// TIA Portal project "Mes_Con" (V17) (continued)
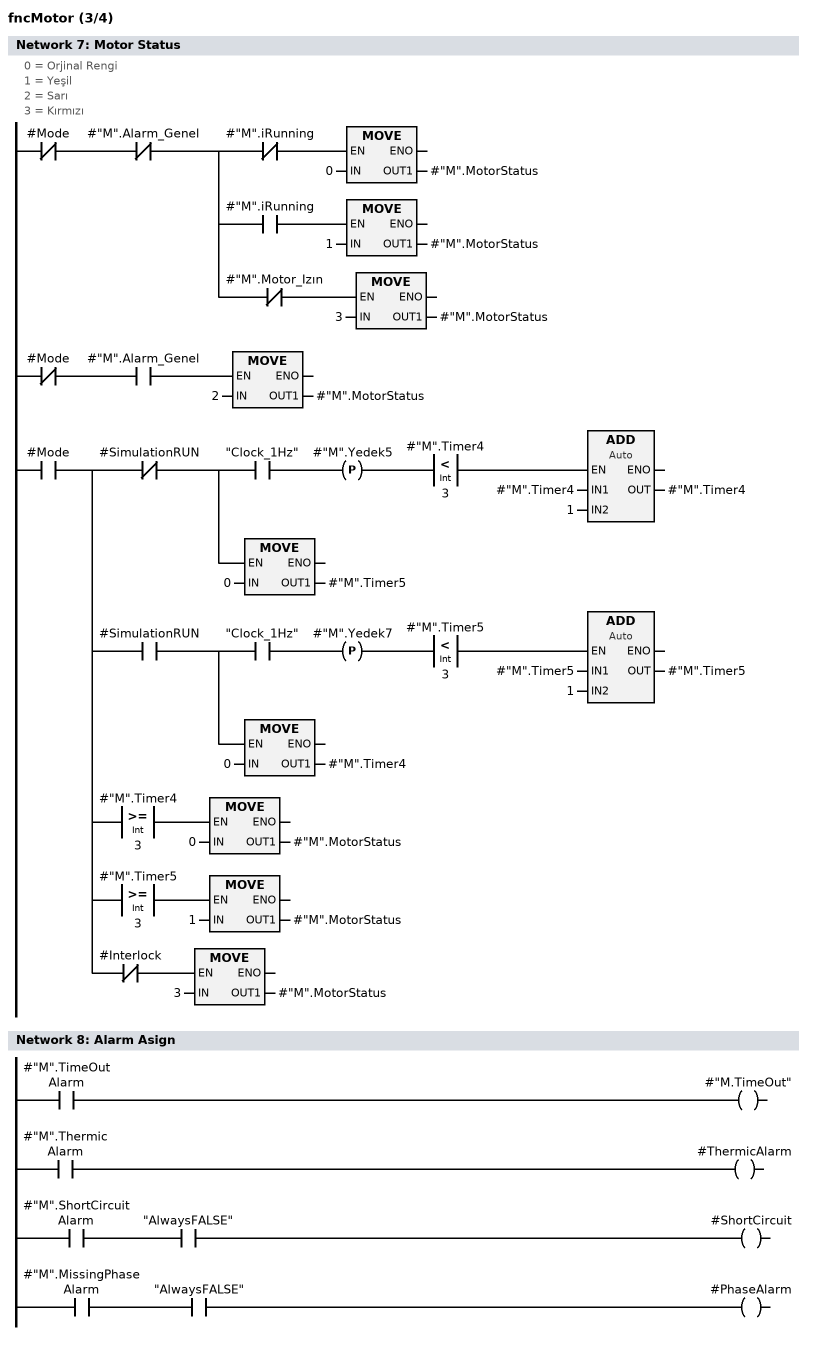
   RUNG wire#powerrail
      I_Contact( #Mode )
      I_Contact( #"M".Alarm_Genel )
      wire#w1
      I_Contact( #"M".iRunning )
      Move(in := 0, out1 => #"M".MotorStatus)
   END_RUNG
   RUNG wire#w1
      Contact( #"M".iRunning )
      Move(in := 1, out1 => #"M".MotorStatus)
   END_RUNG
   RUNG wire#w1
      I_Contact( #"M".Motor_Izın )
      Move(in := 3, out1 => #"M".MotorStatus)
   END_RUNG
   RUNG wire#powerrail
      I_Contact( #Mode )
      Contact( #"M".Alarm_Genel )
      Move(in := 2, out1 => #"M".MotorStatus)
   END_RUNG
   RUNG wire#powerrail
      Contact( #Mode )
      wire#w2
      I_Contact( #SimulationRUN )
      wire#w3
      Contact( "Clock_1Hz" )
      P_Trig( #"M".Yedek5 )
      { S7_Templates := "SrcType := Int" } LT_Contact(in1 := #"M".Timer4, in2 := 3)
      Add(in1 := #"M".Timer4, in2 := 1, out => #"M".Timer4)
   END_RUNG
   RUNG wire#w3
      Move(in := 0, out1 => #"M".Timer5)
   END_RUNG
   RUNG wire#w2
      Contact( #SimulationRUN )
      wire#w4
      Contact( "Clock_1Hz" )
      P_Trig( #"M".Yedek7 )
      { S7_Templates := "SrcType := Int" } LT_Contact(in1 := #"M".Timer5, in2 := 3)
      Add(in1 := #"M".Timer5, in2 := 1, out => #"M".Timer5)
   END_RUNG
   RUNG wire#w4
      Move(in := 0, out1 => #"M".Timer4)
   END_RUNG
   RUNG wire#w2
      { S7_Templates := "SrcType := Int" } GE_Contact(in1 := #"M".Timer4, in2 := 3)
      Move(in := 0, out1 => #"M".MotorStatus)
   END_RUNG
   RUNG wire#w2
      { S7_Templates := "SrcType := Int" } GE_Contact(in1 := #"M".Timer5, in2 := 3)
      Move(in := 1, out1 => #"M".MotorStatus)
   END_RUNG
   RUNG wire#w2
      I_Contact( #Interlock )
      Move(in := 3, out1 => #"M".MotorStatus)
   END_RUNG
   // the same network as SCL:
   #_w1 := NOT #Mode AND NOT #"M".Alarm_Genel;
   IF #_w1 AND NOT #"M".iRunning THEN #"M".MotorStatus := 0; END_IF;
   IF #_w1 AND #"M".iRunning THEN #"M".MotorStatus := 1; END_IF;
   IF #_w1 AND NOT #"M".Motor_Izın THEN #"M".MotorStatus := 3; END_IF;
   IF NOT #Mode AND #"M".Alarm_Genel THEN #"M".MotorStatus := 2; END_IF;
   #_w2 := #Mode AND NOT #SimulationRUN;
   #_w3 := #_w2 AND "Clock_1Hz";
   #_w4 := #_w3 AND NOT #"M".Yedek5;   // rising edge
   #"M".Yedek5 := #_w3;
   IF #_w4 AND (#"M".Timer4 < 3) THEN #"M".Timer4 := #"M".Timer4 + 1; END_IF;
   IF #_w2 THEN #"M".Timer5 := 0; END_IF;
   #_w5 := #Mode AND #SimulationRUN;
   #_w6 := #_w5 AND "Clock_1Hz";
   #_w7 := #_w6 AND NOT #"M".Yedek7;   // rising edge
   #"M".Yedek7 := #_w6;
   IF #_w7 AND (#"M".Timer5 < 3) THEN #"M".Timer5 := #"M".Timer5 + 1; END_IF;
   IF #_w5 THEN #"M".Timer4 := 0; END_IF;
   IF #Mode AND (#"M".Timer4 >= 3) THEN #"M".MotorStatus := 0; END_IF;
   IF #Mode AND (#"M".Timer5 >= 3) THEN #"M".MotorStatus := 1; END_IF;
   IF #Mode AND NOT #Interlock THEN #"M".MotorStatus := 3; END_IF;
END_REGION

REGION Network 8: Alarm Asign
   RUNG wire#powerrail
      Contact( #"M".TimeOutAlarm )
      Coil( #"M.TimeOut" )
   END_RUNG
   RUNG wire#powerrail
      Contact( #"M".ThermicAlarm )
      Coil( #ThermicAlarm )
   END_RUNG
   RUNG wire#powerrail
      Contact( #"M".ShortCircuitAlarm )
      Contact( "AlwaysFALSE" )
      Coil( #ShortCircuit )
   END_RUNG
   RUNG wire#powerrail
      Contact( #"M".MissingPhaseAlarm )
      Contact( "AlwaysFALSE" )
      Coil( #PhaseAlarm )
   END_RUNG
   // the same network as SCL:
   #"M.TimeOut" := #"M".TimeOutAlarm;
   #ThermicAlarm := #"M".ThermicAlarm;
   #ShortCircuit := #"M".ShortCircuitAlarm AND "AlwaysFALSE";
   #PhaseAlarm := #"M".MissingPhaseAlarm AND "AlwaysFALSE";
END_REGION

REGION Network 9: POPUP KAPATMA
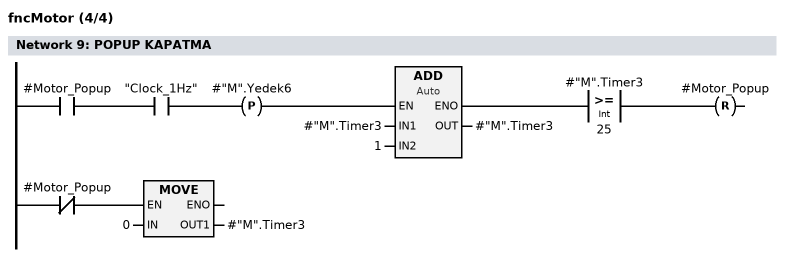
   RUNG wire#powerrail
      Contact( #Motor_Popup )
      Contact( "Clock_1Hz" )
      P_Trig( #"M".Yedek6 )
      Add(in1 := #"M".Timer3, in2 := 1, out => #"M".Timer3)
      { S7_Templates := "SrcType := Int" } GE_Contact(in1 := #"M".Timer3, in2 := 25)
      R_Coil( #Motor_Popup )
   END_RUNG
   RUNG wire#powerrail
      I_Contact( #Motor_Popup )
      Move(in := 0, out1 => #"M".Timer3)
   END_RUNG
   // the same network as SCL:
   #_w1 := #Motor_Popup AND "Clock_1Hz";
   #_w2 := #_w1 AND NOT #"M".Yedek6;   // rising edge
   #"M".Yedek6 := #_w1;
   IF #_w2 THEN #"M".Timer3 := #"M".Timer3 + 1; END_IF;
   IF #_w2 AND (#"M".Timer3 >= 25) THEN #Motor_Popup := FALSE; END_IF;
   IF NOT #Motor_Popup THEN #"M".Timer3 := 0; END_IF;
END_REGION
END_FUNCTION

// folder: Eqp/Valve

FUNCTION "fncValve" : Void   // FC3, LAD
{ S7_Optimized_Access := 'TRUE' }
VERSION : 0.1
   VAR_INPUT
      Mode : Bool;   // 0 = RunTime , 1 = Simulation
      Valve_Opened : Bool;
      Valve_Closed : Bool;
      Interlock : Bool;
   END_VAR
   VAR_OUTPUT
      Valve_Run : Bool;
      Valve_Alarm : Bool;
      Not_Opened : Bool;
      Not_Closed : Bool;
      Not_Signal : Bool;
      Two_Signal : Bool;
   END_VAR
   VAR_IN_OUT
      V : "Valve";
      Vana_Popup : Bool;
   END_VAR
   VAR_TEMP
      SimOpen : Bool;
      SimClose : Bool;
   END_VAR
   VAR_TEMP   // added for the SCL form of the ladder/FBD networks
      _w1 : Bool;
      _w2 : Bool;
      _w3 : Bool;
      _w4 : Bool;
      _w5 : Bool;
      _w6 : Bool;
      _w7 : Bool;
      _w8 : Bool;
      _w9 : Bool;
      _w10 : Bool;
      _w11 : Bool;
      _w12 : Bool;
   END_VAR
BEGIN

REGION Network 1: ATAMA
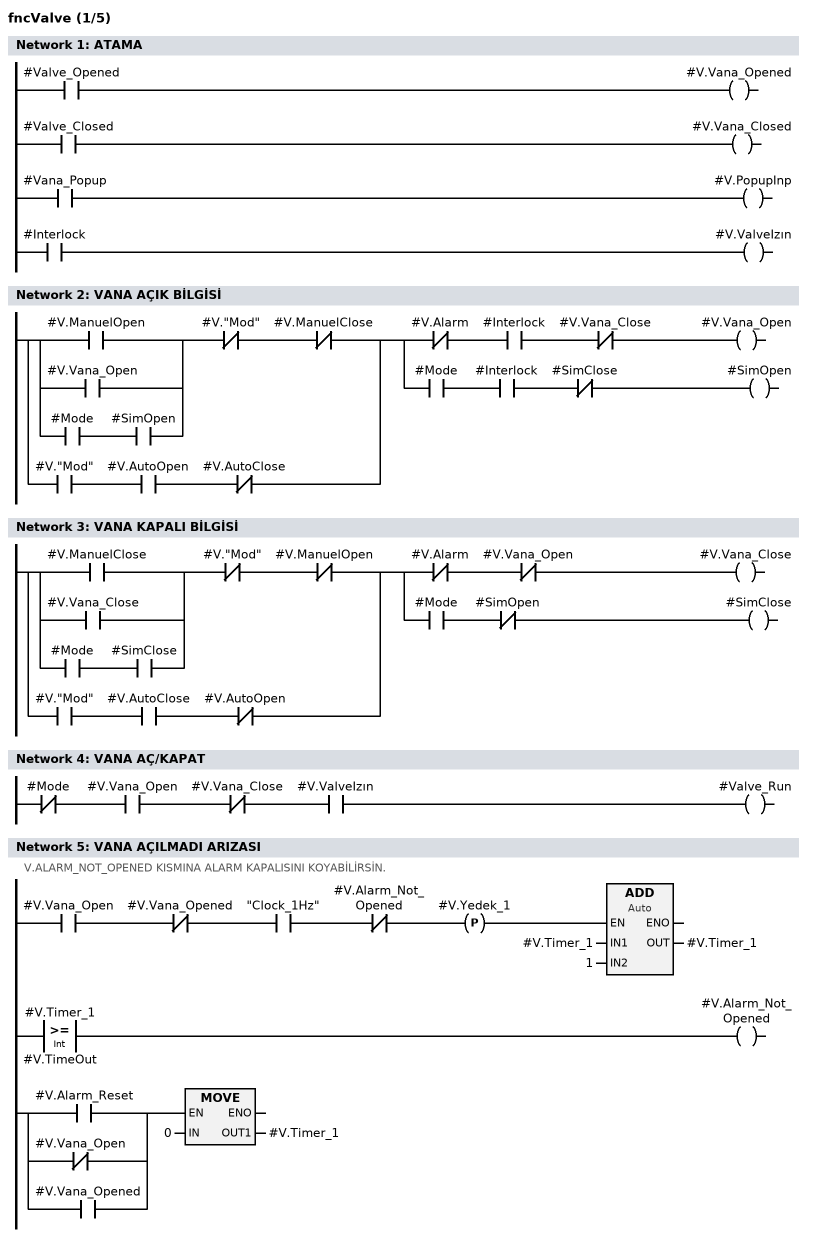
   RUNG wire#powerrail
      Contact( #Valve_Opened )
      Coil( #V.Vana_Opened )
   END_RUNG
   RUNG wire#powerrail
      Contact( #Valve_Closed )
      Coil( #V.Vana_Closed )
   END_RUNG
   RUNG wire#powerrail
      Contact( #Vana_Popup )
      Coil( #V.PopupInp )
   END_RUNG
   RUNG wire#powerrail
      Contact( #Interlock )
      Coil( #V.ValveIzın )
   END_RUNG
   // the same network as SCL:
   #V.Vana_Opened := #Valve_Opened;
   #V.Vana_Closed := #Valve_Closed;
   #V.PopupInp := #Vana_Popup;
   #V.ValveIzın := #Interlock;
END_REGION

REGION Network 2: VANA AÇIK BİLGİSİ
   RUNG wire#powerrail
      Contact( #V.ManuelOpen )
      wire#w1
      I_Contact( #V."Mod" )
      I_Contact( #V.ManuelClose )
      wire#w2
      I_Contact( #V.Alarm )
      Contact( #Interlock )
      I_Contact( #V.Vana_Close )
      Coil( #V.Vana_Open )
   END_RUNG
   RUNG wire#powerrail
      Contact( #V.Vana_Open )
   END_RUNG wire#w1
   RUNG wire#powerrail
      Contact( #Mode )
      Contact( #SimOpen )
   END_RUNG wire#w1
   RUNG wire#powerrail
      Contact( #V."Mod" )
      Contact( #V.AutoOpen )
      I_Contact( #V.AutoClose )
   END_RUNG wire#w2
   RUNG wire#w2
      Contact( #Mode )
      Contact( #Interlock )
      I_Contact( #SimClose )
      Coil( #SimOpen )
   END_RUNG
   // the same network as SCL:
   #_w1 := ((#V.ManuelOpen OR #V.Vana_Open OR (#Mode AND #SimOpen)) AND NOT #V."Mod" AND NOT #V.ManuelClose) OR (#V."Mod" AND #V.AutoOpen AND NOT #V.AutoClose);
   #V.Vana_Open := #_w1 AND NOT #V.Alarm AND #Interlock AND NOT #V.Vana_Close;
   #SimOpen := #_w1 AND #Mode AND #Interlock AND NOT #SimClose;
END_REGION

REGION Network 3: VANA KAPALI BİLGİSİ
   RUNG wire#powerrail
      Contact( #V.ManuelClose )
      wire#w1
      I_Contact( #V."Mod" )
      I_Contact( #V.ManuelOpen )
      wire#w2
      I_Contact( #V.Alarm )
      I_Contact( #V.Vana_Open )
      Coil( #V.Vana_Close )
   END_RUNG
   RUNG wire#powerrail
      Contact( #V.Vana_Close )
   END_RUNG wire#w1
   RUNG wire#powerrail
      Contact( #Mode )
      Contact( #SimClose )
   END_RUNG wire#w1
   RUNG wire#powerrail
      Contact( #V."Mod" )
      Contact( #V.AutoClose )
      I_Contact( #V.AutoOpen )
   END_RUNG wire#w2
   RUNG wire#w2
      Contact( #Mode )
      I_Contact( #SimOpen )
      Coil( #SimClose )
   END_RUNG
   // the same network as SCL:
   #_w1 := ((#V.ManuelClose OR #V.Vana_Close OR (#Mode AND #SimClose)) AND NOT #V."Mod" AND NOT #V.ManuelOpen) OR (#V."Mod" AND #V.AutoClose AND NOT #V.AutoOpen);
   #V.Vana_Close := #_w1 AND NOT #V.Alarm AND NOT #V.Vana_Open;
   #SimClose := #_w1 AND #Mode AND NOT #SimOpen;
END_REGION

REGION Network 4: VANA AÇ/KAPAT
   RUNG wire#powerrail
      I_Contact( #Mode )
      Contact( #V.Vana_Open )
      I_Contact( #V.Vana_Close )
      Contact( #V.ValveIzın )
      Coil( #Valve_Run )
   END_RUNG
   // the same network as SCL:
   #Valve_Run := NOT #Mode AND #V.Vana_Open AND NOT #V.Vana_Close AND #V.ValveIzın;
END_REGION

REGION Network 5: VANA AÇILMADI ARIZASI
   // V.ALARM_NOT_OPENED KISMINA ALARM KAPALISINI KOYABİLİRSİN.
   RUNG wire#powerrail
      Contact( #V.Vana_Open )
      I_Contact( #V.Vana_Opened )
      Contact( "Clock_1Hz" )
      I_Contact( #V.Alarm_Not_Opened )
      P_Trig( #V.Yedek_1 )
      Add(in1 := #V.Timer_1, in2 := 1, out => #V.Timer_1)
   END_RUNG
   RUNG wire#powerrail
      { S7_Templates := "SrcType := Int" } GE_Contact(in1 := #V.Timer_1, in2 := #V.TimeOut)
      Coil( #V.Alarm_Not_Opened )
   END_RUNG
   RUNG wire#powerrail
      Contact( #V.Alarm_Reset )
      wire#w1
      Move(in := 0, out1 => #V.Timer_1)
   END_RUNG
   RUNG wire#powerrail
      I_Contact( #V.Vana_Open )
   END_RUNG wire#w1
   RUNG wire#powerrail
      Contact( #V.Vana_Opened )
   END_RUNG wire#w1
   // the same network as SCL:
   #_w1 := #V.Vana_Open AND NOT #V.Vana_Opened AND "Clock_1Hz" AND NOT #V.Alarm_Not_Opened;
   #_w2 := #_w1 AND NOT #V.Yedek_1;   // rising edge
   #V.Yedek_1 := #_w1;
   IF #_w2 THEN #V.Timer_1 := #V.Timer_1 + 1; END_IF;
   #V.Alarm_Not_Opened := #V.Timer_1 >= #V.TimeOut;
   IF #V.Alarm_Reset OR NOT #V.Vana_Open OR #V.Vana_Opened THEN #V.Timer_1 := 0; END_IF;
END_REGION

REGION Network 6: VANA KAPANMADI ARIZASI
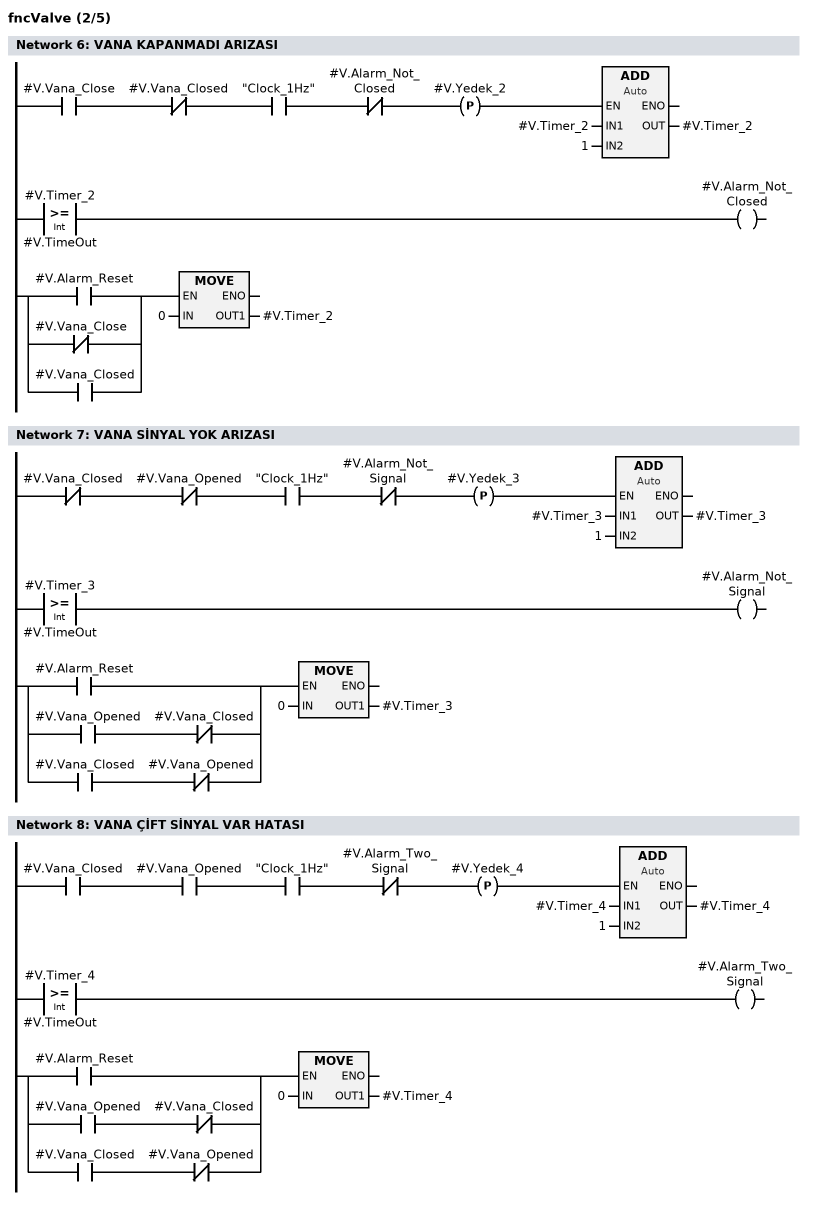
   RUNG wire#powerrail
      Contact( #V.Vana_Close )
      I_Contact( #V.Vana_Closed )
      Contact( "Clock_1Hz" )
      I_Contact( #V.Alarm_Not_Closed )
      P_Trig( #V.Yedek_2 )
      Add(in1 := #V.Timer_2, in2 := 1, out => #V.Timer_2)
   END_RUNG
   RUNG wire#powerrail
      { S7_Templates := "SrcType := Int" } GE_Contact(in1 := #V.Timer_2, in2 := #V.TimeOut)
      Coil( #V.Alarm_Not_Closed )
   END_RUNG
   RUNG wire#powerrail
      Contact( #V.Alarm_Reset )
      wire#w1
      Move(in := 0, out1 => #V.Timer_2)
   END_RUNG
   RUNG wire#powerrail
      I_Contact( #V.Vana_Close )
   END_RUNG wire#w1
   RUNG wire#powerrail
      Contact( #V.Vana_Closed )
   END_RUNG wire#w1
   // the same network as SCL:
   #_w1 := #V.Vana_Close AND NOT #V.Vana_Closed AND "Clock_1Hz" AND NOT #V.Alarm_Not_Closed;
   #_w2 := #_w1 AND NOT #V.Yedek_2;   // rising edge
   #V.Yedek_2 := #_w1;
   IF #_w2 THEN #V.Timer_2 := #V.Timer_2 + 1; END_IF;
   #V.Alarm_Not_Closed := #V.Timer_2 >= #V.TimeOut;
   IF #V.Alarm_Reset OR NOT #V.Vana_Close OR #V.Vana_Closed THEN #V.Timer_2 := 0; END_IF;
END_REGION

REGION Network 7: VANA SİNYAL YOK ARIZASI
   RUNG wire#powerrail
      I_Contact( #V.Vana_Closed )
      I_Contact( #V.Vana_Opened )
      Contact( "Clock_1Hz" )
      I_Contact( #V.Alarm_Not_Signal )
      P_Trig( #V.Yedek_3 )
      Add(in1 := #V.Timer_3, in2 := 1, out => #V.Timer_3)
   END_RUNG
   RUNG wire#powerrail
      { S7_Templates := "SrcType := Int" } GE_Contact(in1 := #V.Timer_3, in2 := #V.TimeOut)
      Coil( #V.Alarm_Not_Signal )
   END_RUNG
   RUNG wire#powerrail
      Contact( #V.Alarm_Reset )
      wire#w1
      Move(in := 0, out1 => #V.Timer_3)
   END_RUNG
   RUNG wire#powerrail
      Contact( #V.Vana_Opened )
      I_Contact( #V.Vana_Closed )
   END_RUNG wire#w1
   RUNG wire#powerrail
      Contact( #V.Vana_Closed )
      I_Contact( #V.Vana_Opened )
   END_RUNG wire#w1
   // the same network as SCL:
   #_w1 := NOT #V.Vana_Closed AND NOT #V.Vana_Opened AND "Clock_1Hz" AND NOT #V.Alarm_Not_Signal;
   #_w2 := #_w1 AND NOT #V.Yedek_3;   // rising edge
   #V.Yedek_3 := #_w1;
   IF #_w2 THEN #V.Timer_3 := #V.Timer_3 + 1; END_IF;
   #V.Alarm_Not_Signal := #V.Timer_3 >= #V.TimeOut;
   IF #V.Alarm_Reset OR (#V.Vana_Opened AND NOT #V.Vana_Closed) OR (#V.Vana_Closed AND NOT #V.Vana_Opened) THEN
       #V.Timer_3 := 0;
   END_IF;
END_REGION

REGION Network 8: VANA ÇİFT SİNYAL VAR HATASI
   RUNG wire#powerrail
      Contact( #V.Vana_Closed )
      Contact( #V.Vana_Opened )
      Contact( "Clock_1Hz" )
      I_Contact( #V.Alarm_Two_Signal )
      P_Trig( #V.Yedek_4 )
      Add(in1 := #V.Timer_4, in2 := 1, out => #V.Timer_4)
   END_RUNG
   RUNG wire#powerrail
      { S7_Templates := "SrcType := Int" } GE_Contact(in1 := #V.Timer_4, in2 := #V.TimeOut)
      Coil( #V.Alarm_Two_Signal )
   END_RUNG
   RUNG wire#powerrail
      Contact( #V.Alarm_Reset )
      wire#w1
      Move(in := 0, out1 => #V.Timer_4)
   END_RUNG
   RUNG wire#powerrail
      Contact( #V.Vana_Opened )
      I_Contact( #V.Vana_Closed )
   END_RUNG wire#w1
   RUNG wire#powerrail
      Contact( #V.Vana_Closed )
      I_Contact( #V.Vana_Opened )
   END_RUNG wire#w1
   // the same network as SCL:
   #_w1 := #V.Vana_Closed AND #V.Vana_Opened AND "Clock_1Hz" AND NOT #V.Alarm_Two_Signal;
   #_w2 := #_w1 AND NOT #V.Yedek_4;   // rising edge
   #V.Yedek_4 := #_w1;
   IF #_w2 THEN #V.Timer_4 := #V.Timer_4 + 1; END_IF;
   #V.Alarm_Two_Signal := #V.Timer_4 >= #V.TimeOut;
   IF #V.Alarm_Reset OR (#V.Vana_Opened AND NOT #V.Vana_Closed) OR (#V.Vana_Closed AND NOT #V.Vana_Opened) THEN
       #V.Timer_4 := 0;
   END_IF;
END_REGION

REGION Network 9: GENEL ALARM
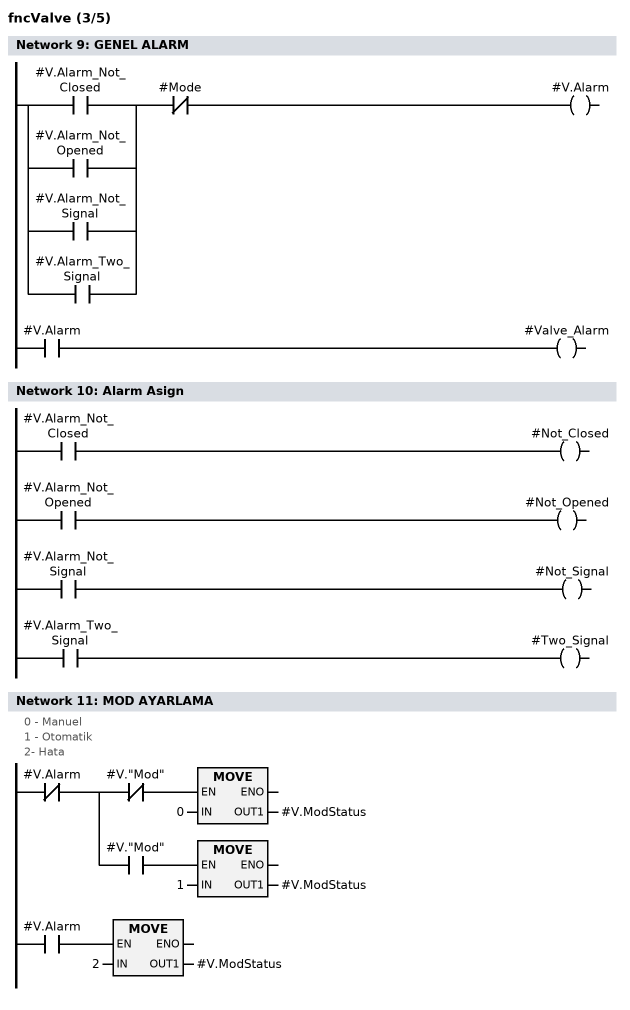
   RUNG wire#powerrail
      Contact( #V.Alarm_Not_Closed )
      wire#w1
      I_Contact( #Mode )
      Coil( #V.Alarm )
   END_RUNG
   RUNG wire#powerrail
      Contact( #V.Alarm_Not_Opened )
   END_RUNG wire#w1
   RUNG wire#powerrail
      Contact( #V.Alarm_Not_Signal )
   END_RUNG wire#w1
   RUNG wire#powerrail
      Contact( #V.Alarm_Two_Signal )
   END_RUNG wire#w1
   RUNG wire#powerrail
      Contact( #V.Alarm )
      Coil( #Valve_Alarm )
   END_RUNG
   // the same network as SCL:
   #V.Alarm := (#V.Alarm_Not_Closed OR #V.Alarm_Not_Opened OR #V.Alarm_Not_Signal OR #V.Alarm_Two_Signal) AND NOT #Mode;
   #Valve_Alarm := #V.Alarm;
END_REGION

REGION Network 10: Alarm Asign
   RUNG wire#powerrail
      Contact( #V.Alarm_Not_Closed )
      Coil( #Not_Closed )
   END_RUNG
   RUNG wire#powerrail
      Contact( #V.Alarm_Not_Opened )
      Coil( #Not_Opened )
   END_RUNG
   RUNG wire#powerrail
      Contact( #V.Alarm_Not_Signal )
      Coil( #Not_Signal )
   END_RUNG
   RUNG wire#powerrail
      Contact( #V.Alarm_Two_Signal )
      Coil( #Two_Signal )
   END_RUNG
   // the same network as SCL:
   #Not_Closed := #V.Alarm_Not_Closed;
   #Not_Opened := #V.Alarm_Not_Opened;
   #Not_Signal := #V.Alarm_Not_Signal;
   #Two_Signal := #V.Alarm_Two_Signal;
END_REGION

REGION Network 11: MOD AYARLAMA
   // 0 - Manuel
   // 1 - Otomatik
   // 2- Hata
   RUNG wire#powerrail
      I_Contact( #V.Alarm )
      wire#w1
      I_Contact( #V."Mod" )
      Move(in := 0, out1 => #V.ModStatus)
   END_RUNG
   RUNG wire#w1
      Contact( #V."Mod" )
      Move(in := 1, out1 => #V.ModStatus)
   END_RUNG
   RUNG wire#powerrail
      Contact( #V.Alarm )
      Move(in := 2, out1 => #V.ModStatus)
   END_RUNG
   // the same network as SCL:
   IF NOT #V.Alarm AND NOT #V."Mod" THEN #V.ModStatus := 0; END_IF;
   IF NOT #V.Alarm AND #V."Mod" THEN #V.ModStatus := 1; END_IF;
   IF #V.Alarm THEN #V.ModStatus := 2; END_IF;
END_REGION

REGION Network 12: STATUS ALMA
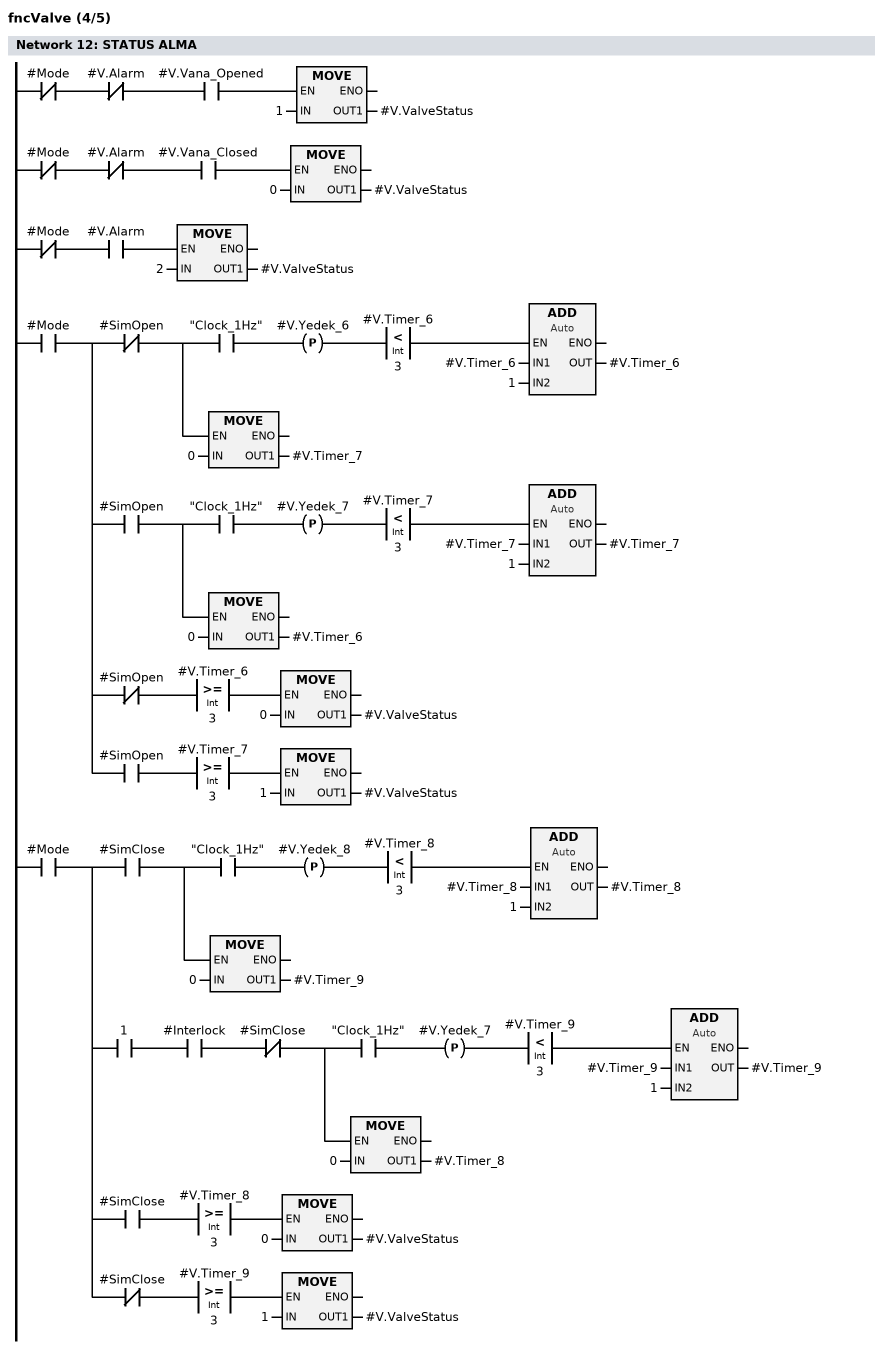
   RUNG wire#powerrail
      I_Contact( #Mode )
      I_Contact( #V.Alarm )
      Contact( #V.Vana_Opened )
      Move(in := 1, out1 => #V.ValveStatus)
   END_RUNG
   RUNG wire#powerrail
      I_Contact( #Mode )
      I_Contact( #V.Alarm )
      Contact( #V.Vana_Closed )
      Move(in := 0, out1 => #V.ValveStatus)
   END_RUNG
   RUNG wire#powerrail
      I_Contact( #Mode )
      Contact( #V.Alarm )
      Move(in := 2, out1 => #V.ValveStatus)
   END_RUNG
   RUNG wire#powerrail
      Contact( #Mode )
      wire#w1
      I_Contact( #SimOpen )
      wire#w2
      Contact( "Clock_1Hz" )
      P_Trig( #V.Yedek_6 )
      { S7_Templates := "SrcType := Int" } LT_Contact(in1 := #V.Timer_6, in2 := 3)
      Add(in1 := #V.Timer_6, in2 := 1, out => #V.Timer_6)
   END_RUNG
   RUNG wire#w2
      Move(in := 0, out1 => #V.Timer_7)
   END_RUNG
   RUNG wire#w1
      Contact( #SimOpen )
      wire#w3
      Contact( "Clock_1Hz" )
      P_Trig( #V.Yedek_7 )
      { S7_Templates := "SrcType := Int" } LT_Contact(in1 := #V.Timer_7, in2 := 3)
      Add(in1 := #V.Timer_7, in2 := 1, out => #V.Timer_7)
   END_RUNG
   RUNG wire#w3
      Move(in := 0, out1 => #V.Timer_6)
   END_RUNG
   RUNG wire#w1
      I_Contact( #SimOpen )
      { S7_Templates := "SrcType := Int" } GE_Contact(in1 := #V.Timer_6, in2 := 3)
      Move(in := 0, out1 => #V.ValveStatus)
   END_RUNG
   RUNG wire#w1
      Contact( #SimOpen )
      { S7_Templates := "SrcType := Int" } GE_Contact(in1 := #V.Timer_7, in2 := 3)
      Move(in := 1, out1 => #V.ValveStatus)
   END_RUNG
   RUNG wire#powerrail
      Contact( #Mode )
      wire#w4
      Contact( #SimClose )
      wire#w5
      Contact( "Clock_1Hz" )
      P_Trig( #V.Yedek_8 )
      { S7_Templates := "SrcType := Int" } LT_Contact(in1 := #V.Timer_8, in2 := 3)
      Add(in1 := #V.Timer_8, in2 := 1, out => #V.Timer_8)
   END_RUNG
   RUNG wire#w5
      Move(in := 0, out1 => #V.Timer_9)
   END_RUNG
   RUNG wire#w4
      Contact( 1 )
      Contact( #Interlock )
      I_Contact( #SimClose )
      wire#w6
      Contact( "Clock_1Hz" )
      P_Trig( #V.Yedek_7 )
      { S7_Templates := "SrcType := Int" } LT_Contact(in1 := #V.Timer_9, in2 := 3)
      Add(in1 := #V.Timer_9, in2 := 1, out => #V.Timer_9)
   END_RUNG
   RUNG wire#w6
      Move(in := 0, out1 => #V.Timer_8)
   END_RUNG
   RUNG wire#w4
      Contact( #SimClose )
      { S7_Templates := "SrcType := Int" } GE_Contact(in1 := #V.Timer_8, in2 := 3)
      Move(in := 0, out1 => #V.ValveStatus)
   END_RUNG
   RUNG wire#w4
      I_Contact( #SimClose )
      { S7_Templates := "SrcType := Int" } GE_Contact(in1 := #V.Timer_9, in2 := 3)
      Move(in := 1, out1 => #V.ValveStatus)
   END_RUNG
   // the same network as SCL:
   IF NOT #Mode AND NOT #V.Alarm AND #V.Vana_Opened THEN #V.ValveStatus := 1; END_IF;
   IF NOT #Mode AND NOT #V.Alarm AND #V.Vana_Closed THEN #V.ValveStatus := 0; END_IF;
   IF NOT #Mode AND #V.Alarm THEN #V.ValveStatus := 2; END_IF;
   #_w1 := #Mode AND NOT #SimOpen;
   #_w2 := #_w1 AND "Clock_1Hz";
   #_w3 := #_w2 AND NOT #V.Yedek_6;   // rising edge
   #V.Yedek_6 := #_w2;
   IF #_w3 AND (#V.Timer_6 < 3) THEN #V.Timer_6 := #V.Timer_6 + 1; END_IF;
   IF #_w1 THEN #V.Timer_7 := 0; END_IF;
   #_w4 := #Mode AND #SimOpen;
   #_w5 := #_w4 AND "Clock_1Hz";
   #_w6 := #_w5 AND NOT #V.Yedek_7;   // rising edge
   #V.Yedek_7 := #_w5;
   IF #_w6 AND (#V.Timer_7 < 3) THEN #V.Timer_7 := #V.Timer_7 + 1; END_IF;
   IF #_w4 THEN #V.Timer_6 := 0; END_IF;
   IF #Mode AND NOT #SimOpen AND (#V.Timer_6 >= 3) THEN #V.ValveStatus := 0; END_IF;
   IF #Mode AND #SimOpen AND (#V.Timer_7 >= 3) THEN #V.ValveStatus := 1; END_IF;
   #_w7 := #Mode AND #SimClose;
   #_w8 := #_w7 AND "Clock_1Hz";
   #_w9 := #_w8 AND NOT #V.Yedek_8;   // rising edge
   #V.Yedek_8 := #_w8;
   IF #_w9 AND (#V.Timer_8 < 3) THEN #V.Timer_8 := #V.Timer_8 + 1; END_IF;
   IF #_w7 THEN #V.Timer_9 := 0; END_IF;
   #_w10 := #Mode AND 1 AND #Interlock AND NOT #SimClose;
   #_w11 := #_w10 AND "Clock_1Hz";
   #_w12 := #_w11 AND NOT #V.Yedek_7;   // rising edge
   #V.Yedek_7 := #_w11;
   IF #_w12 AND (#V.Timer_9 < 3) THEN #V.Timer_9 := #V.Timer_9 + 1; END_IF;
   IF #_w10 THEN #V.Timer_8 := 0; END_IF;
   IF #Mode AND #SimClose AND (#V.Timer_8 >= 3) THEN #V.ValveStatus := 0; END_IF;
   IF #Mode AND NOT #SimClose AND (#V.Timer_9 >= 3) THEN #V.ValveStatus := 1; END_IF;
END_REGION

REGION Network 13: POPUP KAPATMA
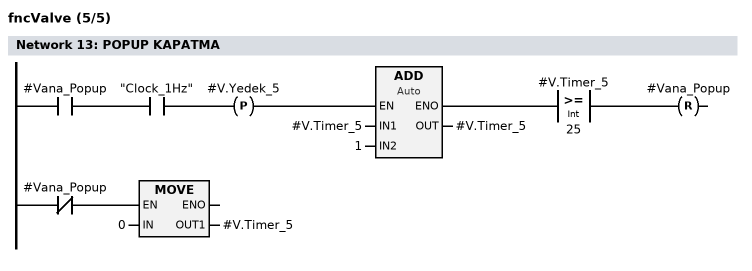
   RUNG wire#powerrail
      Contact( #Vana_Popup )
      Contact( "Clock_1Hz" )
      P_Trig( #V.Yedek_5 )
      Add(in1 := #V.Timer_5, in2 := 1, out => #V.Timer_5)
      { S7_Templates := "SrcType := Int" } GE_Contact(in1 := #V.Timer_5, in2 := 25)
      R_Coil( #Vana_Popup )
   END_RUNG
   RUNG wire#powerrail
      I_Contact( #Vana_Popup )
      Move(in := 0, out1 => #V.Timer_5)
   END_RUNG
   // the same network as SCL:
   #_w1 := #Vana_Popup AND "Clock_1Hz";
   #_w2 := #_w1 AND NOT #V.Yedek_5;   // rising edge
   #V.Yedek_5 := #_w1;
   IF #_w2 THEN #V.Timer_5 := #V.Timer_5 + 1; END_IF;
   IF #_w2 AND (#V.Timer_5 >= 25) THEN #Vana_Popup := FALSE; END_IF;
   IF NOT #Vana_Popup THEN #V.Timer_5 := 0; END_IF;
END_REGION
END_FUNCTION

(* ===== HMI "HMI_RT_1" =====
system functions are stored by id; their names below are inferred from use
connection "HMI_Connection_1": ETHERNET, SMART_S7_1500_OMS

HMI tags "Default tag table"
   "Tag_ScreenNumber" : UInt, internal
   "PUMP_PUMP-1_MotorStatus" : Int = PLC PUMP.PUMP-1.MotorStatus, 1 s
   "PUMP_PUMP-2_MotorStatus" : Int = PLC PUMP.PUMP-2.MotorStatus, 1 s
   "PUMP_PUMP-3_MotorStatus" : Int = PLC PUMP.PUMP-3.MotorStatus, 1 s
   "PUMP_PUMP-4_MotorStatus" : Int = PLC PUMP.PUMP-4.MotorStatus, 1 s
   "VALVE-H_VALVE-1_ValveStatus" : Int = PLC "VALVE-H".VALVE-1.ValveStatus, 1 s
   "VALVE-H_VALVE-2_ValveStatus" : Int = PLC "VALVE-H".VALVE-2.ValveStatus, 1 s
   "VALVE-H_VALVE-3_ValveStatus" : Int = PLC "VALVE-H".VALVE-3.ValveStatus, 1 s
   "VALVE-H_VALVE-4_ValveStatus" : Int = PLC "VALVE-H".VALVE-4.ValveStatus, 1 s
   "Pump-1_Temp" : Word = PLC "Pump-1_Temp" AT %IW124, 1 s
   "Pump-1_A" : Word = PLC "Pump-1_A" AT %IW126, 1 s
   "Pump-2_Temp" : Word = PLC "Pump-2_Temp" AT %IW128, 1 s
   "Pump-2_A" : Word = PLC "Pump-2_A" AT %IW130, 1 s
   "Pump-3_Temp" : Word = PLC "Pump-3_Temp" AT %IW132, 1 s
   "Pump-3_A" : Word = PLC "Pump-3_A" AT %IW134, 1 s
   "Pump-4_Temp" : Word = PLC "Pump-4_Temp" AT %IW136, 1 s
   "Pump-4_A" : Word = PLC "Pump-4_A" AT %IW138, 1 s
   "TT-0001" : Word = PLC "TT-0001" AT %IW116, 1 s
   "TT-0002" : Word = PLC "TT-0002" AT %IW118, 1 s
   "PT-0001" : Word = PLC "PT-0001" AT %IW120, 1 s
   "PT-0002" : Word = PLC "PT-0002" AT %IW122, 1 s
   "CValve-1_Fbk" : Word = PLC "CValve-1_Fbk" AT %IW100, 1 s
   "CValve-2_Fbk" : Word = PLC "CValve-2_Fbk" AT %IW102, 1 s
   "CValve-3_Fbk" : Word = PLC "CValve-3_Fbk" AT %IW104, 1 s
   "CValve-4_Fbk" : Word = PLC "CValve-4_Fbk" AT %IW106, 1 s
   "HMI_Popup_POPUP{8}" : Bool = PLC HMI.Popup.POPUP[8], 1 s
   "HMI_CValve-1_Set" : Int = PLC HMI.CValve-1_Set, 1 s
   "HMI_Popup_POPUP{9}" : Bool = PLC HMI.Popup.POPUP[9], 1 s
   "HMI_CValve-2_Set" : Int = PLC HMI.CValve-2_Set, 1 s
   "HMI_Popup_POPUP{10}" : Bool = PLC HMI.Popup.POPUP[10], 1 s
   "HMI_CValve-3_Set" : Int = PLC HMI.CValve-3_Set, 1 s
   "HMI_Popup_POPUP{11}" : Bool = PLC HMI.Popup.POPUP[11], 1 s
   "HMI_Popup_POPUP{0}" : Bool = PLC HMI.Popup.POPUP[0], 1 s
   "PUMP_PUMP-1_ManuelStart" : Bool = PLC PUMP.PUMP-1.ManuelStart, 1 s
   "PUMP_PUMP-1_ManuelStop" : Bool = PLC PUMP.PUMP-1.ManuelStop, 1 s
   "HMI_Pump-1" : Int = PLC HMI.Pump-1, 1 s
   "HMI_Popup_POPUP{1}" : Bool = PLC HMI.Popup.POPUP[1], 1 s
   "PUMP_PUMP-2_ManuelStart" : Bool = PLC PUMP.PUMP-2.ManuelStart, 1 s
   "PUMP_PUMP-2_ManuelStop" : Bool = PLC PUMP.PUMP-2.ManuelStop, 1 s
   "HMI_Pump-2" : Int = PLC HMI.Pump-2, 1 s
   "HMI_Popup_POPUP{2}" : Bool = PLC HMI.Popup.POPUP[2], 1 s
   "PUMP_PUMP-3_ManuelStart" : Bool = PLC PUMP.PUMP-3.ManuelStart, 1 s
   "PUMP_PUMP-3_ManuelStop" : Bool = PLC PUMP.PUMP-3.ManuelStop, 1 s
   "HMI_Popup_POPUP{3}" : Bool = PLC HMI.Popup.POPUP[3], 1 s
   "HMI_Pump-3" : Int = PLC HMI.Pump-3, 1 s
   "HMI_Pump-4" : Int = PLC HMI.Pump-4, 1 s
   "PUMP_PUMP-4_ManuelStart" : Bool = PLC PUMP.PUMP-4.ManuelStart, 1 s
   "PUMP_PUMP-4_ManuelStop" : Bool = PLC PUMP.PUMP-4.ManuelStop, 1 s
   "PUMP_PUMP-1_Local/Remote" : Bool = PLC PUMP.PUMP-1.Local/Remote, 1 s
   "PUMP_PUMP-2_Local/Remote" : Bool = PLC PUMP.PUMP-2.Local/Remote, 1 s
   "PUMP_PUMP-3_Local/Remote" : Bool = PLC PUMP.PUMP-3.Local/Remote, 1 s
   "PUMP_PUMP-4_Local/Remote" : Bool = PLC PUMP.PUMP-4.Local/Remote, 1 s
   "HMI_Popup_POPUP{4}" : Bool = PLC HMI.Popup.POPUP[4], 1 s
   "VALVE-H_VALVE-1_Vana_Opened" : Bool = PLC "VALVE-H".VALVE-1.Vana_Opened, 1 s
   "VALVE-H_VALVE-1_ManuelOpen" : Bool = PLC "VALVE-H".VALVE-1.ManuelOpen, 1 s
   "HMI_Popup_POPUP{5}" : Bool = PLC HMI.Popup.POPUP[5], 1 s
   "HMI_Popup_POPUP{6}" : Bool = PLC HMI.Popup.POPUP[6], 1 s
   "HMI_Popup_POPUP{7}" : Bool = PLC HMI.Popup.POPUP[7], 1 s
   "VALVE-H_VALVE-2_Vana_Opened" : Bool = PLC "VALVE-H".VALVE-2.Vana_Opened, 1 s
   "VALVE-H_VALVE-3_Vana_Opened" : Bool = PLC "VALVE-H".VALVE-3.Vana_Opened, 1 s
   "VALVE-H_VALVE-4_Vana_Opened" : Bool = PLC "VALVE-H".VALVE-4.Vana_Opened, 1 s
   "VALVE-H_VALVE-2_ManuelOpen" : Bool = PLC "VALVE-H".VALVE-2.ManuelOpen, 1 s
   "VALVE-H_VALVE-3_ManuelClose" : Bool = PLC "VALVE-H".VALVE-3.ManuelClose, 1 s
   "VALVE-H_VALVE-3_ManuelOpen" : Bool = PLC "VALVE-H".VALVE-3.ManuelOpen, 1 s
   "VALVE-H_VALVE-4_ManuelOpen" : Bool = PLC "VALVE-H".VALVE-4.ManuelOpen, 1 s
   "Sim_SİM_MOD" : Bool = PLC Sim.SİM_MOD, 1 s
   "VALVE-H_VALVE-4_ManuelClose" : Bool = PLC "VALVE-H".VALVE-4.ManuelClose, 1 s
   "VALVE-H_VALVE-1_ManuelClose" : Bool = PLC "VALVE-H".VALVE-1.ManuelClose, 1 s
   "VALVE-H_VALVE-2_ManuelClose" : Bool = PLC "VALVE-H".VALVE-2.ManuelClose, 1 s
   "Sim_SPUMP-1_Thermic" : Bool = PLC Sim.SPUMP-1_Thermic, 1 s
   "Sim_SPUMP-2_Thermic" : Bool = PLC Sim.SPUMP-2_Thermic, 1 s
   "Sim_SPUMP-3_Thermic" : Bool = PLC Sim.SPUMP-3_Thermic, 1 s
   "Sim_SPUMP-4_Thermic" : Bool = PLC Sim.SPUMP-4_Thermic, 1 s
   "Sim_SPUMP-1_Loc" : Bool = PLC Sim.SPUMP-1_Loc, 1 s
   "Sim_SPUMP-2_Loc" : Bool = PLC Sim.SPUMP-2_Loc, 1 s
   "Sim_SPUMP-3_Loc" : Bool = PLC Sim.SPUMP-3_Loc, 1 s
   "Sim_SPUMP-4_Loc" : Bool = PLC Sim.SPUMP-4_Loc, 1 s
   "Sim_SPump-1_RPM" : Word = PLC Sim.SPump-1_RPM, 1 s
   "Sim_SPump-2_RPM" : Word = PLC Sim.SPump-2_RPM, 1 s
   "Sim_SPump-3_RPM" : Word = PLC Sim.SPump-3_RPM, 1 s
   "Sim_SPump-4_RPM" : Word = PLC Sim.SPump-4_RPM, 1 s
   "Sim_SPump-1_Temp" : Word = PLC Sim.SPump-1_Temp, 1 s
   "Sim_SPump-2_Temp" : Word = PLC Sim.SPump-2_Temp, 1 s
   "Sim_SPump-3_Temp" : Word = PLC Sim.SPump-3_Temp, 1 s
   "Sim_SPump-4_Temp" : Word = PLC Sim.SPump-4_Temp, 1 s
   "Sim_SPump-1_A" : Word = PLC Sim.SPump-1_A, 1 s
   "Sim_SPump-2_A" : Word = PLC Sim.SPump-2_A, 1 s
   "Sim_SPump-3_A" : Word = PLC Sim.SPump-3_A, 1 s
   "Sim_SPump-4_A" : Word = PLC Sim.SPump-4_A, 1 s
   "Sim_SCValve-1_Fbk" : Word = PLC Sim.SCValve-1_Fbk, 1 s
   "Sim_SCValve-2_Fbk" : Word = PLC Sim.SCValve-2_Fbk, 1 s
   "Sim_SCValve-3_Fbk" : Word = PLC Sim.SCValve-3_Fbk, 1 s
   "Sim_SCValve-4_Fbk" : Word = PLC Sim.SCValve-4_Fbk, 1 s
   "Sim_STT-0001" : Word = PLC Sim.STT-0001, 1 s
   "Sim_STT-0002" : Word = PLC Sim.STT-0002, 1 s
   "Sim_SPT-0001" : Word = PLC Sim.SPT-0001, 1 s
   "Sim_SPT-0002" : Word = PLC Sim.SPT-0002, 1 s
   "workorder_Work_Order-1_Active" : Bool = PLC workorder.Work_Order-1_Active AT %DB10.DBX0.0, 1 s
   "workorder_Work_Order-2_Active" : Bool = PLC workorder.Work_Order-2_Active AT %DB10.DBX0.1, 1 s
   "workorder_Work_Order-3_Active" : Bool = PLC workorder.Work_Order-3_Active AT %DB10.DBX0.2, 1 s
   "workorder_Work_Order-4_Active" : Bool = PLC workorder.Work_Order-4_Active AT %DB10.DBX0.3, 1 s
   "workorder_Work_Order-5_Active" : Bool = PLC workorder.Work_Order-5_Active AT %DB10.DBX0.4, 1 s
   "workorder_Work_Order-6_Active" : Bool = PLC workorder.Work_Order-6_Active AT %DB10.DBX0.5, 1 s
   "workorder_Work_Order-7_Active" : Bool = PLC workorder.Work_Order-7_Active AT %DB10.DBX0.6, 1 s
   "workorder_Work_Order-8_Active" : Bool = PLC workorder.Work_Order-8_Active AT %DB10.DBX0.7, 1 s
   "workorder_Work_Order-9_Active" : Bool = PLC workorder.Work_Order-9_Active AT %DB10.DBX1.0, 1 s
   "workorder_Work_Order-10_Active" : Bool = PLC workorder.Work_Order-10_Active AT %DB10.DBX1.1, 1 s
   "workorder_Work_Order-11_Active" : Bool = PLC workorder.Work_Order-11_Active AT %DB10.DBX1.2, 1 s
   "workorder_Work_Order-12_Active" : Bool = PLC workorder.Work_Order-12_Active AT %DB10.DBX1.3, 1 s
   "workorder_Work_Order-13_Active" : Bool = PLC workorder.Work_Order-13_Active AT %DB10.DBX1.4, 1 s
   "workorder_Work_Order-14_Active" : Bool = PLC workorder.Work_Order-14_Active AT %DB10.DBX1.5, 1 s
   "PUMP-1_Loc" : Bool = PLC "PUMP-1_Loc" AT %I10.2, 1 s
   "PUMP_PUMP-1_Yedek1" : Bool = PLC PUMP.PUMP-1.Yedek1, 1 s
   "PUMP_PUMP-2_Yedek1" : Bool = PLC PUMP.PUMP-2.Yedek1, 1 s
   "PUMP_PUMP-3_Yedek1" : Bool = PLC PUMP.PUMP-3.Yedek1, 1 s
   "PUMP_PUMP-4_Yedek1" : Bool = PLC PUMP.PUMP-4.Yedek1, 1 s
   "HMI_CValve-4_Set" : Int = PLC HMI.CValve-4_Set, 1 s

text list "Kullanici_Tanimla": 2 'Operatör'; 3 'Yönetici'; 1 'İzleyici'; 4 'Tanker Mod'

text list "WorkOrder": 1 'Work Order-1'; 2 'Work Order-2'; 3 'Work Order-3'; 4 'Work Order-4'; 5 'Work Order-5'; 6 'Work Order-6'; 7 'Work Order-7'; 8 'Work Order-8'; 9 'Work Order-9'; 10 'Work Order-10'; 11 'Work Order-11'; 12 'Work Order-12'; 13 'Work Order-13'; 14 'Work Order-14'

Template "Template_1" 800x480
   DateTimeField "HmiScreenItemData" at 714,29 size 80x20
      ProcessValue <- "TARİH_SAAT__YEREL_SAAT"
   DateTimeField "HmiScreenItemData_1" at 722,7 size 71x20
      ProcessValue <- "TARİH_SAAT__YEREL_SAAT"
   Button "Button_12" at 19,9 size 241x43; TextOff 'ANA SAYFA'
   Button "Template_Button_1" at 283,8 size 60x47; TextOff 'Text'; PictureOff "home-button_1"
      on Press: ActivateScreen("Proses", 0)
   Button "Template_Button_2" at 366,8 size 60x47; TextOff 'Text'; PictureOff "generative"
      on Press: ActivateScreen("Con", 0)
   Button "Template_Button_3" at 443,8 size 60x47; TextOff 'Text'; PictureOff "done_3"
      on Press: ActivateScreen("todolist", 0)
   Button "Template_Button_4" at 584,7 size 60x47; TextOff 'Text'; PictureOff "alert_2"
   Button "Template_Button_5" at 654,7 size 60x47; TextOff 'Text'; PictureOff "profile_2"
   Button "Template_Button_6" at 515,8 size 60x47; TextOff 'Text'; PictureOff "simulation"
      on Press: ActivateScreen("simkontrol", 0)

screen "dd" 800x480, template "Template_1"
   on GenerateScreen: SetTag("Tag_ScreenNumber", 1)

screen "simkontrol" 800x480, template "Template_1"
   Switch "Switch_6" at 100,65 size 120x34; TextOn 'ON'; CaptionText 'Switch'; TextOff 'OFF'
      ProcessValue <- "Sim_SİM_MOD"
   TextField "Text field_6" at 14,71 size 74x20; Text 'Sim Status'
   TextField "Text field_1" at 80,126 size 61x20; Text 'THERMIC'
   TextField "Text field_2" at 14,152 size 54x20; Text 'PUMP-1'
   TextField "Text field_3" at 14,202 size 54x20; Text 'PUMP-2'
   TextField "Text field_4" at 14,251 size 54x20; Text 'PUMP-3'
   TextField "Text field_5" at 14,298 size 54x20; Text 'PUMP-4'
   TextField "Text field_7" at 170,124 size 46x20; Text 'LOCAL'
   Switch "Switch_1" at 160,144 size 80x35; TextOn 'ON'; CaptionText 'Switch'; TextOff 'OFF'
      ProcessValue <- "Sim_SPUMP-1_Loc"
   Switch "Switch_2" at 160,194 size 80x35; TextOn 'ON'; CaptionText 'Switch'; TextOff 'OFF'
      ProcessValue <- "Sim_SPUMP-2_Loc"
   Switch "Switch_3" at 160,243 size 80x35; TextOn 'ON'; CaptionText 'Switch'; TextOff 'OFF'
      ProcessValue <- "Sim_SPUMP-3_Loc"
   Switch "Switch_4" at 160,290 size 80x35; TextOn 'ON'; CaptionText 'Switch'; TextOff 'OFF'
      ProcessValue <- "Sim_SPUMP-4_Loc"
   Switch "Switch_5" at 78,144 size 80x35; TextOn 'ON'; CaptionText 'Switch'; TextOff 'OFF'
      ProcessValue <- "Sim_SPUMP-1_Thermic"
   Switch "Switch_7" at 78,194 size 80x35; TextOn 'ON'; CaptionText 'Switch'; TextOff 'OFF'
      ProcessValue <- "Sim_SPUMP-2_Thermic"
   Switch "Switch_8" at 78,243 size 80x35; TextOn 'ON'; CaptionText 'Switch'; TextOff 'OFF'
      ProcessValue <- "Sim_SPUMP-3_Thermic"
   Switch "Switch_9" at 78,290 size 80x35; TextOn 'ON'; CaptionText 'Switch'; TextOff 'OFF'
      ProcessValue <- "Sim_SPUMP-4_Thermic"
   TextField "Text field_8" at 255,128 size 33x20; Text 'RPM'
   TextField "Text field_9" at 334,128 size 42x20; Text 'TEMP.'
   TextField "Text field_10" at 395,128 size 15x20; Text 'A'
   IOField "I/O field_11" at 326,152 size 60x26; FormatPattern 999; Unit  °C
      ProcessValue <- "Sim_SPump-1_Temp"
   IOField "I/O field_5" at 395,152 size 49x26; FormatPattern 99; Unit  A
      ProcessValue <- "Sim_SPump-1_A"
   IOField "I/O field_1" at 245,152 size 69x26; FormatPattern 999; Unit  rpm
      ProcessValue <- "Sim_SPump-1_RPM"
   IOField "I/O field_2" at 326,202 size 60x26; FormatPattern 999; Unit  °C
      ProcessValue <- "Sim_SPump-2_Temp"
   IOField "I/O field_3" at 395,202 size 49x26; FormatPattern 99; Unit  A
      ProcessValue <- "Sim_SPump-2_A"
   IOField "I/O field_4" at 245,202 size 69x26; FormatPattern 999; Unit  rpm
      ProcessValue <- "Sim_SPump-2_RPM"
   IOField "I/O field_6" at 326,251 size 60x26; FormatPattern 999; Unit  °C
      ProcessValue <- "Sim_SPump-3_Temp"
   IOField "I/O field_7" at 395,251 size 49x26; FormatPattern 99; Unit  A
      ProcessValue <- "Sim_SPump-3_A"
   IOField "I/O field_8" at 245,251 size 69x26; FormatPattern 999; Unit  rpm
      ProcessValue <- "Sim_SPump-3_RPM"
   IOField "I/O field_9" at 326,298 size 60x26; FormatPattern 999; Unit  °C
      ProcessValue <- "Sim_SPump-4_Temp"
   IOField "I/O field_10" at 395,298 size 49x26; FormatPattern 99; Unit  A
      ProcessValue <- "Sim_SPump-4_A"
   IOField "I/O field_12" at 245,298 size 69x26; FormatPattern 999; Unit  rpm
      ProcessValue <- "Sim_SPump-4_RPM"
   TextField "Text field_11" at 472,258 size 67x20; Text 'C.Valve-1'
   TextField "Text field_12" at 472,289 size 67x20; Text 'C.Valve-2'
   TextField "Text field_13" at 472,320 size 67x20; Text 'C.Valve-3'
   TextField "Text field_14" at 472,352 size 67x20; Text 'C.Valve-4'
   IOField "I/O field_13" at 558,258 size 65x20; FormatPattern 999; Unit  %
      ProcessValue <- "Sim_SCValve-1_Fbk"
   IOField "I/O field_14" at 558,289 size 65x20; FormatPattern 999; Unit  %
      ProcessValue <- "Sim_SCValve-2_Fbk"
   IOField "I/O field_15" at 558,320 size 65x20; FormatPattern 999; Unit  %
      ProcessValue <- "Sim_SCValve-3_Fbk"
   IOField "I/O field_16" at 558,352 size 65x20; FormatPattern 999; Unit  %
      ProcessValue <- "Sim_SCValve-4_Fbk"
   TextField "Text field_15" at 472,115 size 57x20; Text 'TT-0001'
   TextField "Text field_16" at 472,146 size 57x20; Text 'TT-0002'
   TextField "Text field_17" at 472,177 size 58x20; Text 'PT-0001'
   TextField "Text field_18" at 472,209 size 58x20; Text 'PT-0002'
   IOField "I/O field_17" at 558,115 size 56x20; FormatPattern 999; Unit  °C
      ProcessValue <- "Sim_STT-0001"
   IOField "I/O field_18" at 558,146 size 56x20; FormatPattern 999; Unit  °C
      ProcessValue <- "Sim_STT-0002"
   IOField "I/O field_19" at 558,177 size 56x20; FormatPattern 99; Unit  Bar
      ProcessValue <- "Sim_SPT-0001"
   IOField "I/O field_20" at 558,209 size 56x20; FormatPattern 99; Unit  Bar
      ProcessValue <- "Sim_SPT-0002"

